// TIA Portal project "Automatizare_RT" (V17) (continued)
REGION Network 14: Cand sistemul hidraulic este in eroare / Wenn das Hydrauliksystem fehlerhaft ist
   RUNG wire#powerrail
      I_Contact( "DB_general".CondOptimePistoane )
      wire#w1
      { S7_GenerateENO := "TRUE" } Move(in := 0, out1 => "DB_Status_Pistoane".Status_Piston_1)
   END_RUNG
   RUNG wire#w1
      { S7_GenerateENO := "TRUE" } Move(in := 0, out1 => "DB_Status_Pistoane".Status_Pison_2)
   END_RUNG
   RUNG wire#w1
      { S7_GenerateENO := "TRUE" } Move(in := 0, out1 => "DB_Status_Pistoane".Status_Piston_A)
   END_RUNG
   RUNG wire#w1
      { S7_GenerateENO := "TRUE" } Move(in := 0, out1 => "DB_Status_Pistoane".Status_Piston_B)
   END_RUNG
   RUNG wire#w1
      { S7_GenerateENO := "TRUE" } Move(in := 0, out1 => "DB_Status_Pistoane".Status_Piston_C)
   END_RUNG
   // the same network as SCL:
   IF NOT "DB_general".CondOptimePistoane THEN
       "DB_Status_Pistoane".Status_Piston_1 := 0;
       "DB_Status_Pistoane".Status_Pison_2 := 0;
       "DB_Status_Pistoane".Status_Piston_A := 0;
       "DB_Status_Pistoane".Status_Piston_B := 0;
       "DB_Status_Pistoane".Status_Piston_C := 0;
   END_IF;
END_REGION
END_FUNCTION

FUNCTION "Status_Motoare" : Void   // FC8, LAD
{ S7_Optimized_Access := 'FALSE' }
VERSION : 0.1
BEGIN

REGION Network 1: motor 1/2 e in functiune
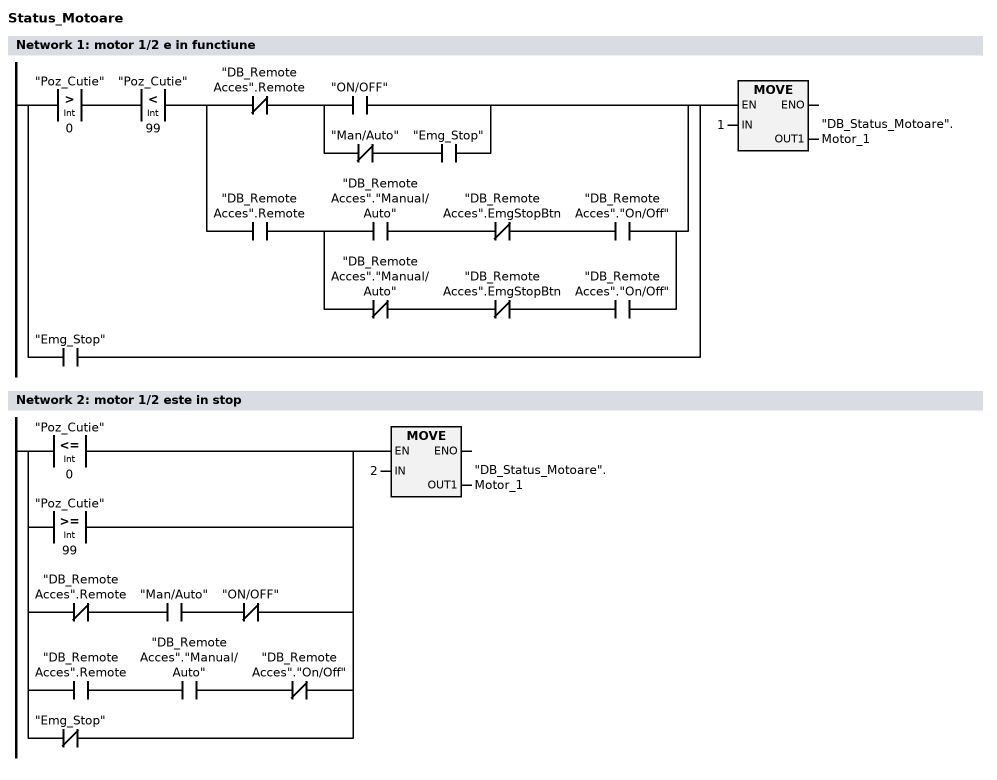
   RUNG wire#powerrail
      { S7_Templates := "SrcType := Int" } GT_Contact(in1 := "Poz_Cutie", in2 := 0)
      { S7_Templates := "SrcType := Int" } LT_Contact(in1 := "Poz_Cutie", in2 := 99)
      wire#w1
      I_Contact( "DB_RemoteAcces".Remote )
      wire#w2
      Contact( "ON/OFF" )
      wire#w3
      { S7_GenerateENO := "TRUE" } Move(in := 1, out1 => "DB_Status_Motoare".Motor_1)
   END_RUNG
   RUNG wire#w2
      I_Contact( "Man/Auto" )
      Contact( "Emg_Stop" )
   END_RUNG wire#w3
   RUNG wire#w1
      Contact( "DB_RemoteAcces".Remote )
      wire#w4
      Contact( "DB_RemoteAcces"."Manual/Auto" )
      I_Contact( "DB_RemoteAcces".EmgStopBtn )
      Contact( "DB_RemoteAcces"."On/Off" )
   END_RUNG wire#w3
   RUNG wire#w4
      I_Contact( "DB_RemoteAcces"."Manual/Auto" )
      I_Contact( "DB_RemoteAcces".EmgStopBtn )
      Contact( "DB_RemoteAcces"."On/Off" )
   END_RUNG wire#w3
   RUNG wire#powerrail
      Contact( "Emg_Stop" )
   END_RUNG wire#w3
   // the same network as SCL:
   IF (("Poz_Cutie" > 0) AND ("Poz_Cutie" < 99) AND ((NOT "DB_RemoteAcces".Remote AND ("ON/OFF" OR (NOT "Man/Auto" AND "Emg_Stop"))) OR ("DB_RemoteAcces".Remote AND (("DB_RemoteAcces"."Manual/Auto" AND NOT "DB_RemoteAcces".EmgStopBtn AND "DB_RemoteAcces"."On/Off") OR (NOT "DB_RemoteAcces"."Manual/Auto" AND NOT "DB_RemoteAcces".EmgStopBtn AND "DB_RemoteAcces"."On/Off"))))) OR "Emg_Stop" THEN
       "DB_Status_Motoare".Motor_1 := 1;
   END_IF;
END_REGION

REGION Network 2: motor 1/2 este in stop
   RUNG wire#powerrail
      { S7_Templates := "SrcType := Int" } LE_Contact(in1 := "Poz_Cutie", in2 := 0)
      wire#w1
      { S7_GenerateENO := "TRUE" } Move(in := 2, out1 => "DB_Status_Motoare".Motor_1)
   END_RUNG
   RUNG wire#powerrail
      { S7_Templates := "SrcType := Int" } GE_Contact(in1 := "Poz_Cutie", in2 := 99)
   END_RUNG wire#w1
   RUNG wire#powerrail
      I_Contact( "DB_RemoteAcces".Remote )
      Contact( "Man/Auto" )
      I_Contact( "ON/OFF" )
   END_RUNG wire#w1
   RUNG wire#powerrail
      Contact( "DB_RemoteAcces".Remote )
      Contact( "DB_RemoteAcces"."Manual/Auto" )
      I_Contact( "DB_RemoteAcces"."On/Off" )
   END_RUNG wire#w1
   RUNG wire#powerrail
      I_Contact( "Emg_Stop" )
   END_RUNG wire#w1
   // the same network as SCL:
   IF ("Poz_Cutie" <= 0) OR ("Poz_Cutie" >= 99) OR (NOT "DB_RemoteAcces".Remote AND "Man/Auto" AND NOT "ON/OFF") OR ("DB_RemoteAcces".Remote AND "DB_RemoteAcces"."Manual/Auto" AND NOT "DB_RemoteAcces"."On/Off") OR NOT "Emg_Stop" THEN
       "DB_Status_Motoare".Motor_1 := 2;
   END_IF;
END_REGION
END_FUNCTION

FUNCTION "CantarFcn" : Void   // FC10, LAD
{ S7_Optimized_Access := 'FALSE' }
VERSION : 0.1
BEGIN

REGION Network 1
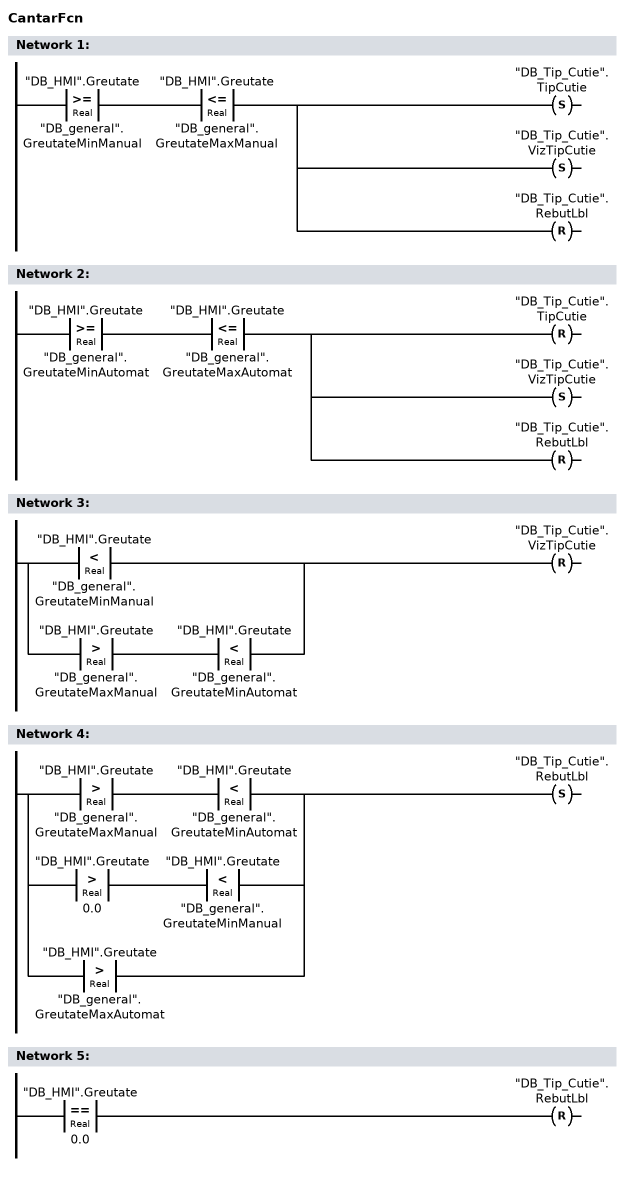
   RUNG wire#powerrail
      { S7_Templates := "SrcType := Real" } GE_Contact(in1 := "DB_HMI".Greutate, in2 := "DB_general".GreutateMinManual)
      { S7_Templates := "SrcType := Real" } LE_Contact(in1 := "DB_HMI".Greutate, in2 := "DB_general".GreutateMaxManual)
      wire#w1
      S_Coil( "DB_Tip_Cutie".TipCutie )
   END_RUNG
   RUNG wire#w1
      S_Coil( "DB_Tip_Cutie".VizTipCutie )
   END_RUNG
   RUNG wire#w1
      R_Coil( "DB_Tip_Cutie".RebutLbl )
   END_RUNG
   // the same network as SCL:
   IF ("DB_HMI".Greutate >= "DB_general".GreutateMinManual) AND ("DB_HMI".Greutate <= "DB_general".GreutateMaxManual) THEN
       "DB_Tip_Cutie".TipCutie := TRUE;
       "DB_Tip_Cutie".VizTipCutie := TRUE;
       "DB_Tip_Cutie".RebutLbl := FALSE;
   END_IF;
END_REGION

REGION Network 2
   RUNG wire#powerrail
      { S7_Templates := "SrcType := Real" } GE_Contact(in1 := "DB_HMI".Greutate, in2 := "DB_general".GreutateMinAutomat)
      { S7_Templates := "SrcType := Real" } LE_Contact(in1 := "DB_HMI".Greutate, in2 := "DB_general".GreutateMaxAutomat)
      wire#w1
      R_Coil( "DB_Tip_Cutie".TipCutie )
   END_RUNG
   RUNG wire#w1
      S_Coil( "DB_Tip_Cutie".VizTipCutie )
   END_RUNG
   RUNG wire#w1
      R_Coil( "DB_Tip_Cutie".RebutLbl )
   END_RUNG
   // the same network as SCL:
   IF ("DB_HMI".Greutate >= "DB_general".GreutateMinAutomat) AND ("DB_HMI".Greutate <= "DB_general".GreutateMaxAutomat) THEN
       "DB_Tip_Cutie".TipCutie := FALSE;
       "DB_Tip_Cutie".VizTipCutie := TRUE;
       "DB_Tip_Cutie".RebutLbl := FALSE;
   END_IF;
END_REGION

REGION Network 3
   RUNG wire#powerrail
      { S7_Templates := "SrcType := Real" } LT_Contact(in1 := "DB_HMI".Greutate, in2 := "DB_general".GreutateMinManual)
      wire#w1
      R_Coil( "DB_Tip_Cutie".VizTipCutie )
   END_RUNG
   RUNG wire#powerrail
      { S7_Templates := "SrcType := Real" } GT_Contact(in1 := "DB_HMI".Greutate, in2 := "DB_general".GreutateMaxManual)
      { S7_Templates := "SrcType := Real" } LT_Contact(in1 := "DB_HMI".Greutate, in2 := "DB_general".GreutateMinAutomat)
   END_RUNG wire#w1
   // the same network as SCL:
   IF ("DB_HMI".Greutate < "DB_general".GreutateMinManual) OR (("DB_HMI".Greutate > "DB_general".GreutateMaxManual) AND ("DB_HMI".Greutate < "DB_general".GreutateMinAutomat)) THEN
       "DB_Tip_Cutie".VizTipCutie := FALSE;
   END_IF;
END_REGION

REGION Network 4
   RUNG wire#powerrail
      { S7_Templates := "SrcType := Real" } GT_Contact(in1 := "DB_HMI".Greutate, in2 := "DB_general".GreutateMaxManual)
      { S7_Templates := "SrcType := Real" } LT_Contact(in1 := "DB_HMI".Greutate, in2 := "DB_general".GreutateMinAutomat)
      wire#w1
      S_Coil( "DB_Tip_Cutie".RebutLbl )
   END_RUNG
   RUNG wire#powerrail
      { S7_Templates := "SrcType := Real" } GT_Contact(in1 := "DB_HMI".Greutate, in2 := 0.0)
      { S7_Templates := "SrcType := Real" } LT_Contact(in1 := "DB_HMI".Greutate, in2 := "DB_general".GreutateMinManual)
   END_RUNG wire#w1
   RUNG wire#powerrail
      { S7_Templates := "SrcType := Real" } GT_Contact(in1 := "DB_HMI".Greutate, in2 := "DB_general".GreutateMaxAutomat)
   END_RUNG wire#w1
   // the same network as SCL:
   IF (("DB_HMI".Greutate > "DB_general".GreutateMaxManual) AND ("DB_HMI".Greutate < "DB_general".GreutateMinAutomat)) OR (("DB_HMI".Greutate > 0.0) AND ("DB_HMI".Greutate < "DB_general".GreutateMinManual)) OR ("DB_HMI".Greutate > "DB_general".GreutateMaxAutomat) THEN
       "DB_Tip_Cutie".RebutLbl := TRUE;
   END_IF;
END_REGION

REGION Network 5
   RUNG wire#powerrail
      { S7_Templates := "SrcType := Real" } EQ_Contact(in1 := "DB_HMI".Greutate, in2 := 0.0)
      R_Coil( "DB_Tip_Cutie".RebutLbl )
   END_RUNG
   // the same network as SCL:
   IF "DB_HMI".Greutate = 0.0 THEN "DB_Tip_Cutie".RebutLbl := FALSE; END_IF;
END_REGION
END_FUNCTION

FUNCTION "CondOptimePistoane" : Void   // FC11, LAD
{ S7_Optimized_Access := 'FALSE' }
VERSION : 0.1
BEGIN

REGION Network 1
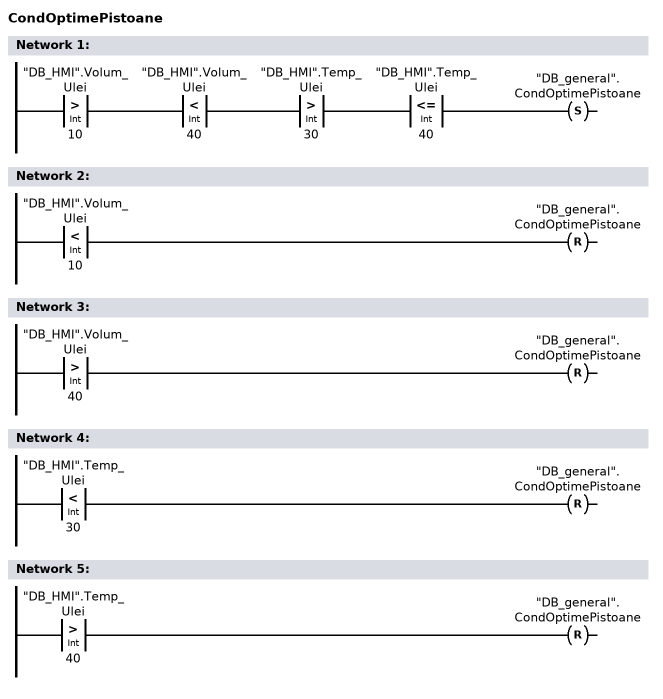
   RUNG wire#powerrail
      { S7_Templates := "SrcType := Int" } GT_Contact(in1 := "DB_HMI".Volum_Ulei, in2 := 10)
      { S7_Templates := "SrcType := Int" } LT_Contact(in1 := "DB_HMI".Volum_Ulei, in2 := 40)
      { S7_Templates := "SrcType := Int" } GT_Contact(in1 := "DB_HMI".Temp_Ulei, in2 := 30)
      { S7_Templates := "SrcType := Int" } LE_Contact(in1 := "DB_HMI".Temp_Ulei, in2 := 40)
      S_Coil( "DB_general".CondOptimePistoane )
   END_RUNG
   // the same network as SCL:
   IF ("DB_HMI".Volum_Ulei > 10) AND ("DB_HMI".Volum_Ulei < 40) AND ("DB_HMI".Temp_Ulei > 30) AND ("DB_HMI".Temp_Ulei <= 40) THEN
       "DB_general".CondOptimePistoane := TRUE;
   END_IF;
END_REGION

REGION Network 2
   RUNG wire#powerrail
      { S7_Templates := "SrcType := Int" } LT_Contact(in1 := "DB_HMI".Volum_Ulei, in2 := 10)
      R_Coil( "DB_general".CondOptimePistoane )
   END_RUNG
   // the same network as SCL:
   IF "DB_HMI".Volum_Ulei < 10 THEN "DB_general".CondOptimePistoane := FALSE; END_IF;
END_REGION

REGION Network 3
   RUNG wire#powerrail
      { S7_Templates := "SrcType := Int" } GT_Contact(in1 := "DB_HMI".Volum_Ulei, in2 := 40)
      R_Coil( "DB_general".CondOptimePistoane )
   END_RUNG
   // the same network as SCL:
   IF "DB_HMI".Volum_Ulei > 40 THEN "DB_general".CondOptimePistoane := FALSE; END_IF;
END_REGION

REGION Network 4
   RUNG wire#powerrail
      { S7_Templates := "SrcType := Int" } LT_Contact(in1 := "DB_HMI".Temp_Ulei, in2 := 30)
      R_Coil( "DB_general".CondOptimePistoane )
   END_RUNG
   // the same network as SCL:
   IF "DB_HMI".Temp_Ulei < 30 THEN "DB_general".CondOptimePistoane := FALSE; END_IF;
END_REGION

REGION Network 5
   RUNG wire#powerrail
      { S7_Templates := "SrcType := Int" } GT_Contact(in1 := "DB_HMI".Temp_Ulei, in2 := 40)
      R_Coil( "DB_general".CondOptimePistoane )
   END_RUNG
   // the same network as SCL:
   IF "DB_HMI".Temp_Ulei > 40 THEN "DB_general".CondOptimePistoane := FALSE; END_IF;
END_REGION
END_FUNCTION

FUNCTION "EroareIntervaleGreutate" : Void   // FC15, STL
{ S7_Optimized_Access := 'FALSE' }
VERSION : 0.1
BEGIN

REGION Network 1


         L     "DB_general".GreutateManual;
         L     "DB_general".Procent_Toleranta;
         *D;
         L     100;
         /R;
         T     "DB_general".TolerantaManual;
         L     "DB_general".TolerantaManual;
         L     "DB_general".GreutateManual;
         +R;
         T     "DB_general".TolerantaManual;
END_REGION
END_FUNCTION

FUNCTION "TipCutieTranzit" : Void   // FC16, LAD
{ S7_Optimized_Access := 'FALSE' }
VERSION : 0.1
BEGIN

REGION Network 1
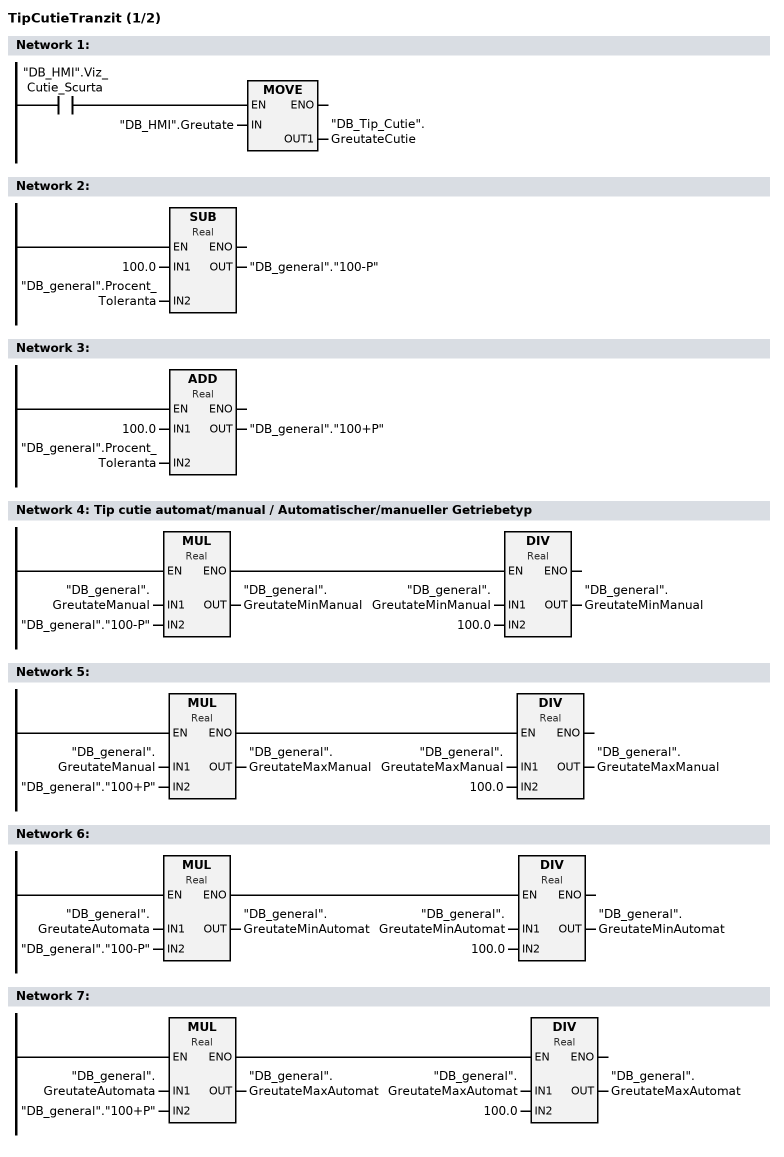
   RUNG wire#powerrail
      Contact( "DB_HMI".Viz_Cutie_Scurta )
      { S7_GenerateENO := "TRUE" } Move(in := "DB_HMI".Greutate, out1 => "DB_Tip_Cutie".GreutateCutie)
   END_RUNG
   // the same network as SCL:
   IF "DB_HMI".Viz_Cutie_Scurta THEN "DB_Tip_Cutie".GreutateCutie := "DB_HMI".Greutate; END_IF;
END_REGION

REGION Network 2
   RUNG wire#powerrail
      { S7_Templates := "SrcType := Real"; S7_GenerateENO := "TRUE" } Sub(in1 := 100.0, in2 := "DB_general".Procent_Toleranta, out => "DB_general"."100-P")
   END_RUNG
   // the same network as SCL:
   "DB_general"."100-P" := 100.0 - "DB_general".Procent_Toleranta;
END_REGION

REGION Network 3
   RUNG wire#powerrail
      { S7_Templates := "SrcType := Real"; S7_GenerateENO := "TRUE" } Add(in1 := 100.0, in2 := "DB_general".Procent_Toleranta, out => "DB_general"."100+P")
   END_RUNG
   // the same network as SCL:
   "DB_general"."100+P" := 100.0 + "DB_general".Procent_Toleranta;
END_REGION

REGION Network 4: Tip cutie automat/manual / Automatischer/manueller Getriebetyp
   RUNG wire#powerrail
      { S7_Templates := "SrcType := Real"; S7_GenerateENO := "TRUE" } Mul(in1 := "DB_general".GreutateManual, in2 := "DB_general"."100-P", out => "DB_general".GreutateMinManual)
      { S7_Templates := "SrcType := Real"; S7_GenerateENO := "TRUE" } Div(in1 := "DB_general".GreutateMinManual, in2 := 100.0, out => "DB_general".GreutateMinManual)
   END_RUNG
   // the same network as SCL:
   // ENO of a box is taken as its EN; it also drops when the box reports an error
   "DB_general".GreutateMinManual := "DB_general".GreutateManual * "DB_general"."100-P";
   "DB_general".GreutateMinManual := "DB_general".GreutateMinManual / 100.0;
END_REGION

REGION Network 5
   RUNG wire#powerrail
      { S7_Templates := "SrcType := Real"; S7_GenerateENO := "TRUE" } Mul(in1 := "DB_general".GreutateManual, in2 := "DB_general"."100+P", out => "DB_general".GreutateMaxManual)
      { S7_Templates := "SrcType := Real"; S7_GenerateENO := "TRUE" } Div(in1 := "DB_general".GreutateMaxManual, in2 := 100.0, out => "DB_general".GreutateMaxManual)
   END_RUNG
   // the same network as SCL:
   // ENO of a box is taken as its EN; it also drops when the box reports an error
   "DB_general".GreutateMaxManual := "DB_general".GreutateManual * "DB_general"."100+P";
   "DB_general".GreutateMaxManual := "DB_general".GreutateMaxManual / 100.0;
END_REGION

REGION Network 6
   RUNG wire#powerrail
      { S7_Templates := "SrcType := Real"; S7_GenerateENO := "TRUE" } Mul(in1 := "DB_general".GreutateAutomata, in2 := "DB_general"."100-P", out => "DB_general".GreutateMinAutomat)
      { S7_Templates := "SrcType := Real"; S7_GenerateENO := "TRUE" } Div(in1 := "DB_general".GreutateMinAutomat, in2 := 100.0, out => "DB_general".GreutateMinAutomat)
   END_RUNG
   // the same network as SCL:
   // ENO of a box is taken as its EN; it also drops when the box reports an error
   "DB_general".GreutateMinAutomat := "DB_general".GreutateAutomata * "DB_general"."100-P";
   "DB_general".GreutateMinAutomat := "DB_general".GreutateMinAutomat / 100.0;
END_REGION

REGION Network 7
   RUNG wire#powerrail
      { S7_Templates := "SrcType := Real"; S7_GenerateENO := "TRUE" } Mul(in1 := "DB_general".GreutateAutomata, in2 := "DB_general"."100+P", out => "DB_general".GreutateMaxAutomat)
      { S7_Templates := "SrcType := Real"; S7_GenerateENO := "TRUE" } Div(in1 := "DB_general".GreutateMaxAutomat, in2 := 100.0, out => "DB_general".GreutateMaxAutomat)
   END_RUNG
   // the same network as SCL:
   // ENO of a box is taken as its EN; it also drops when the box reports an error
   "DB_general".GreutateMaxAutomat := "DB_general".GreutateAutomata * "DB_general"."100+P";
   "DB_general".GreutateMaxAutomat := "DB_general".GreutateMaxAutomat / 100.0;
END_REGION

REGION Network 8
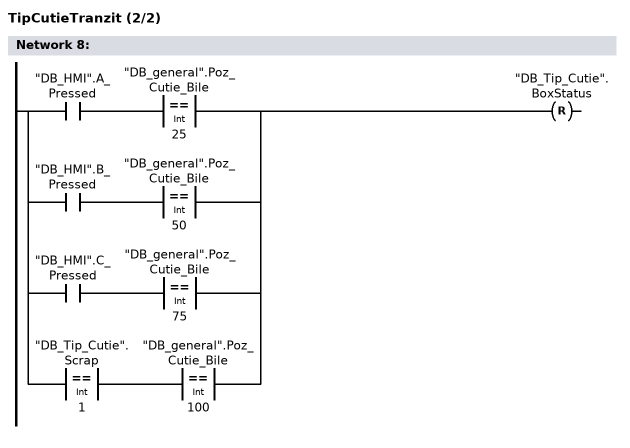
   RUNG wire#powerrail
      Contact( "DB_HMI".A_Pressed )
      { S7_Templates := "SrcType := Int" } EQ_Contact(in1 := "DB_general".Poz_Cutie_Bile, in2 := 25)
      wire#w1
      R_Coil( "DB_Tip_Cutie".BoxStatus )
   END_RUNG
   RUNG wire#powerrail
      Contact( "DB_HMI".B_Pressed )
      { S7_Templates := "SrcType := Int" } EQ_Contact(in1 := "DB_general".Poz_Cutie_Bile, in2 := 50)
   END_RUNG wire#w1
   RUNG wire#powerrail
      Contact( "DB_HMI".C_Pressed )
      { S7_Templates := "SrcType := Int" } EQ_Contact(in1 := "DB_general".Poz_Cutie_Bile, in2 := 75)
   END_RUNG wire#w1
   RUNG wire#powerrail
      { S7_Templates := "SrcType := Int" } EQ_Contact(in1 := "DB_Tip_Cutie".Scrap, in2 := 1)
      { S7_Templates := "SrcType := Int" } EQ_Contact(in1 := "DB_general".Poz_Cutie_Bile, in2 := 100)
   END_RUNG wire#w1
   // the same network as SCL:
   IF ("DB_HMI".A_Pressed AND ("DB_general".Poz_Cutie_Bile = 25)) OR ("DB_HMI".B_Pressed AND ("DB_general".Poz_Cutie_Bile = 50)) OR ("DB_HMI".C_Pressed AND ("DB_general".Poz_Cutie_Bile = 75)) OR (("DB_Tip_Cutie".Scrap = 1) AND ("DB_general".Poz_Cutie_Bile = 100)) THEN
       "DB_Tip_Cutie".BoxStatus := FALSE;
   END_IF;
END_REGION
END_FUNCTION

FUNCTION "EroriCantarire" : Void   // FC17, LAD
{ S7_Optimized_Access := 'FALSE' }
VERSION : 0.1
BEGIN

REGION Network 1
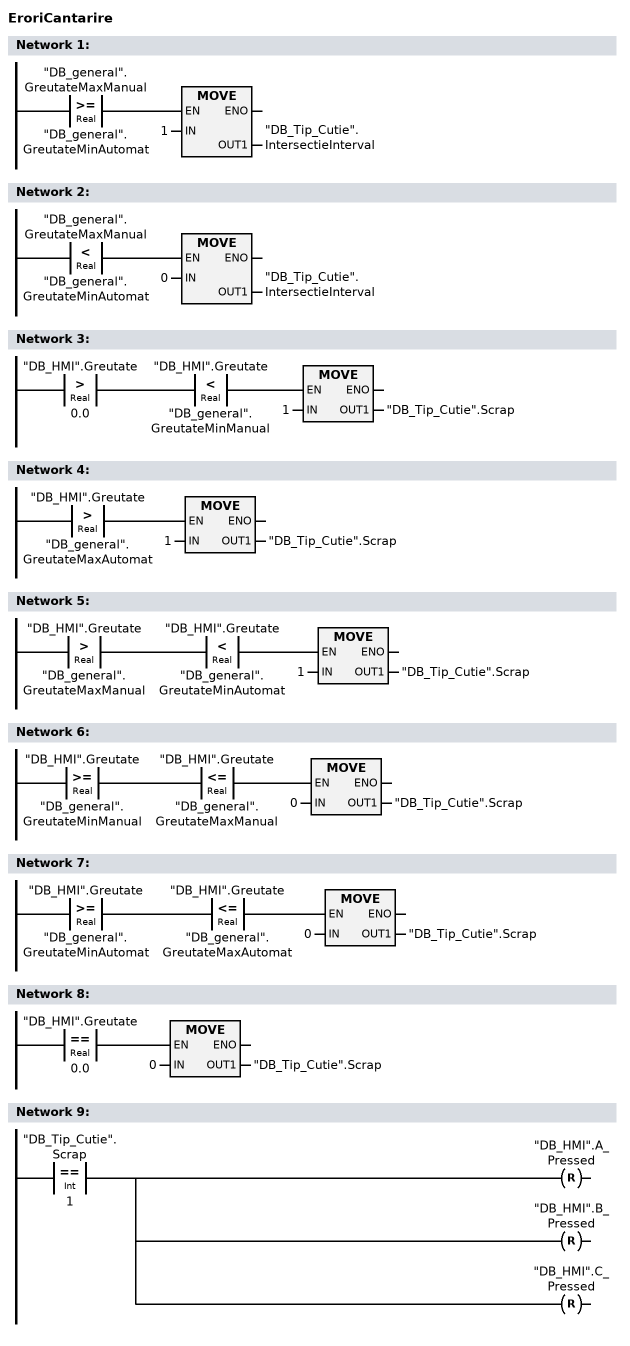
   RUNG wire#powerrail
      { S7_Templates := "SrcType := Real" } GE_Contact(in1 := "DB_general".GreutateMaxManual, in2 := "DB_general".GreutateMinAutomat)
      { S7_GenerateENO := "TRUE" } Move(in := 1, out1 => "DB_Tip_Cutie".IntersectieInterval)
   END_RUNG
   // the same network as SCL:
   IF "DB_general".GreutateMaxManual >= "DB_general".GreutateMinAutomat THEN
       "DB_Tip_Cutie".IntersectieInterval := 1;
   END_IF;
END_REGION

REGION Network 2
   RUNG wire#powerrail
      { S7_Templates := "SrcType := Real" } LT_Contact(in1 := "DB_general".GreutateMaxManual, in2 := "DB_general".GreutateMinAutomat)
      { S7_GenerateENO := "TRUE" } Move(in := 0, out1 => "DB_Tip_Cutie".IntersectieInterval)
   END_RUNG
   // the same network as SCL:
   IF "DB_general".GreutateMaxManual < "DB_general".GreutateMinAutomat THEN
       "DB_Tip_Cutie".IntersectieInterval := 0;
   END_IF;
END_REGION

REGION Network 3
   RUNG wire#powerrail
      { S7_Templates := "SrcType := Real" } GT_Contact(in1 := "DB_HMI".Greutate, in2 := 0.0)
      { S7_Templates := "SrcType := Real" } LT_Contact(in1 := "DB_HMI".Greutate, in2 := "DB_general".GreutateMinManual)
      { S7_GenerateENO := "TRUE" } Move(in := 1, out1 => "DB_Tip_Cutie".Scrap)
   END_RUNG
   // the same network as SCL:
   IF ("DB_HMI".Greutate > 0.0) AND ("DB_HMI".Greutate < "DB_general".GreutateMinManual) THEN
       "DB_Tip_Cutie".Scrap := 1;
   END_IF;
END_REGION

REGION Network 4
   RUNG wire#powerrail
      { S7_Templates := "SrcType := Real" } GT_Contact(in1 := "DB_HMI".Greutate, in2 := "DB_general".GreutateMaxAutomat)
      { S7_GenerateENO := "TRUE" } Move(in := 1, out1 => "DB_Tip_Cutie".Scrap)
   END_RUNG
   // the same network as SCL:
   IF "DB_HMI".Greutate > "DB_general".GreutateMaxAutomat THEN "DB_Tip_Cutie".Scrap := 1; END_IF;
END_REGION

REGION Network 5
   RUNG wire#powerrail
      { S7_Templates := "SrcType := Real" } GT_Contact(in1 := "DB_HMI".Greutate, in2 := "DB_general".GreutateMaxManual)
      { S7_Templates := "SrcType := Real" } LT_Contact(in1 := "DB_HMI".Greutate, in2 := "DB_general".GreutateMinAutomat)
      { S7_GenerateENO := "TRUE" } Move(in := 1, out1 => "DB_Tip_Cutie".Scrap)
   END_RUNG
   // the same network as SCL:
   IF ("DB_HMI".Greutate > "DB_general".GreutateMaxManual) AND ("DB_HMI".Greutate < "DB_general".GreutateMinAutomat) THEN
       "DB_Tip_Cutie".Scrap := 1;
   END_IF;
END_REGION

REGION Network 6
   RUNG wire#powerrail
      { S7_Templates := "SrcType := Real" } GE_Contact(in1 := "DB_HMI".Greutate, in2 := "DB_general".GreutateMinManual)
      { S7_Templates := "SrcType := Real" } LE_Contact(in1 := "DB_HMI".Greutate, in2 := "DB_general".GreutateMaxManual)
      { S7_GenerateENO := "TRUE" } Move(in := 0, out1 => "DB_Tip_Cutie".Scrap)
   END_RUNG
   // the same network as SCL:
   IF ("DB_HMI".Greutate >= "DB_general".GreutateMinManual) AND ("DB_HMI".Greutate <= "DB_general".GreutateMaxManual) THEN
       "DB_Tip_Cutie".Scrap := 0;
   END_IF;
END_REGION

REGION Network 7
   RUNG wire#powerrail
      { S7_Templates := "SrcType := Real" } GE_Contact(in1 := "DB_HMI".Greutate, in2 := "DB_general".GreutateMinAutomat)
      { S7_Templates := "SrcType := Real" } LE_Contact(in1 := "DB_HMI".Greutate, in2 := "DB_general".GreutateMaxAutomat)
      { S7_GenerateENO := "TRUE" } Move(in := 0, out1 => "DB_Tip_Cutie".Scrap)
   END_RUNG
   // the same network as SCL:
   IF ("DB_HMI".Greutate >= "DB_general".GreutateMinAutomat) AND ("DB_HMI".Greutate <= "DB_general".GreutateMaxAutomat) THEN
       "DB_Tip_Cutie".Scrap := 0;
   END_IF;
END_REGION

REGION Network 8
   RUNG wire#powerrail
      { S7_Templates := "SrcType := Real" } EQ_Contact(in1 := "DB_HMI".Greutate, in2 := 0.0)
      { S7_GenerateENO := "TRUE" } Move(in := 0, out1 => "DB_Tip_Cutie".Scrap)
   END_RUNG
   // the same network as SCL:
   IF "DB_HMI".Greutate = 0.0 THEN "DB_Tip_Cutie".Scrap := 0; END_IF;
END_REGION

REGION Network 9
   RUNG wire#powerrail
      { S7_Templates := "SrcType := Int" } EQ_Contact(in1 := "DB_Tip_Cutie".Scrap, in2 := 1)
      wire#w1
      R_Coil( "DB_HMI".A_Pressed )
   END_RUNG
   RUNG wire#w1
      R_Coil( "DB_HMI".B_Pressed )
   END_RUNG
   RUNG wire#w1
      R_Coil( "DB_HMI".C_Pressed )
   END_RUNG
   // the same network as SCL:
   IF "DB_Tip_Cutie".Scrap = 1 THEN
       "DB_HMI".A_Pressed := FALSE;
       "DB_HMI".B_Pressed := FALSE;
       "DB_HMI".C_Pressed := FALSE;
   END_IF;
END_REGION
END_FUNCTION

FUNCTION "ConsolaComanda" : Void   // FC21, LAD
{ S7_Optimized_Access := 'FALSE' }
VERSION : 0.1
   VAR_TEMP   // added for the SCL form of the ladder/FBD networks
      _w1 : Bool;
   END_VAR
BEGIN

REGION Network 1
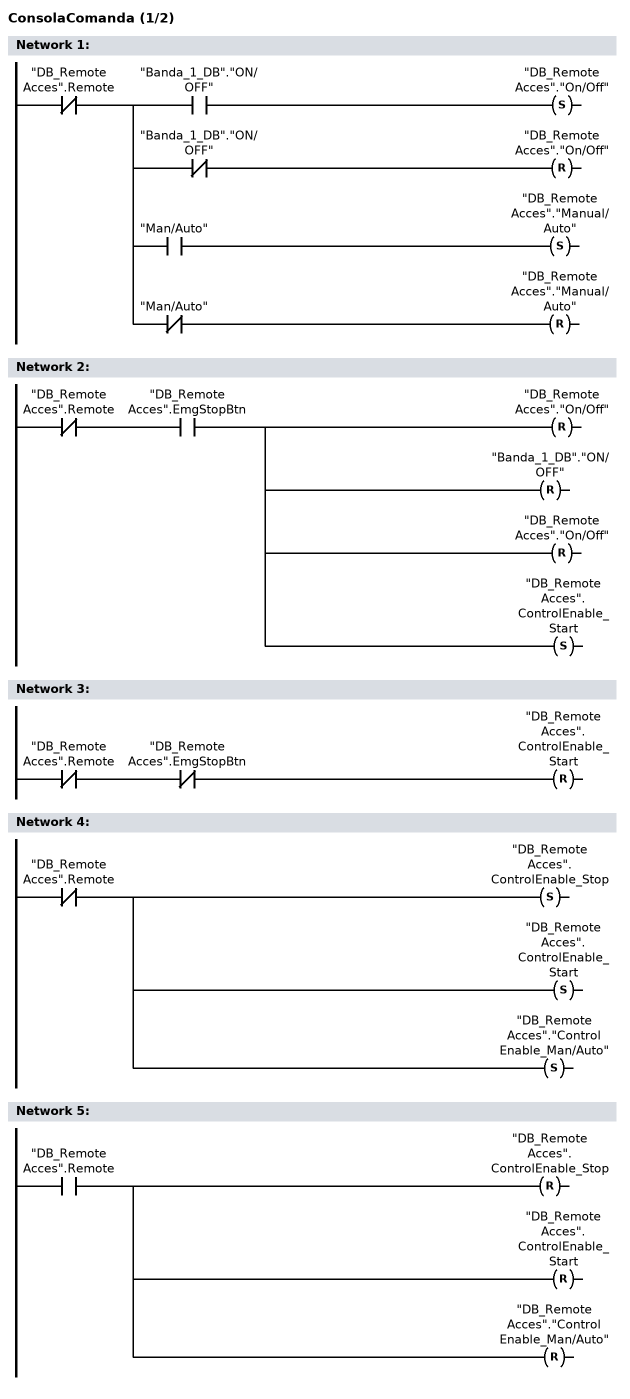
   RUNG wire#powerrail
      I_Contact( "DB_RemoteAcces".Remote )
      wire#w1
      Contact( "Banda_1_DB"."ON/OFF" )
      S_Coil( "DB_RemoteAcces"."On/Off" )
   END_RUNG
   RUNG wire#w1
      I_Contact( "Banda_1_DB"."ON/OFF" )
      R_Coil( "DB_RemoteAcces"."On/Off" )
   END_RUNG
   RUNG wire#w1
      Contact( "Man/Auto" )
      S_Coil( "DB_RemoteAcces"."Manual/Auto" )
   END_RUNG
   RUNG wire#w1
      I_Contact( "Man/Auto" )
      R_Coil( "DB_RemoteAcces"."Manual/Auto" )
   END_RUNG
   // the same network as SCL:
   #_w1 := NOT "DB_RemoteAcces".Remote;
   IF #_w1 AND "Banda_1_DB"."ON/OFF" THEN "DB_RemoteAcces"."On/Off" := TRUE; END_IF;
   IF #_w1 AND NOT "Banda_1_DB"."ON/OFF" THEN "DB_RemoteAcces"."On/Off" := FALSE; END_IF;
   IF #_w1 AND "Man/Auto" THEN "DB_RemoteAcces"."Manual/Auto" := TRUE; END_IF;
   IF #_w1 AND NOT "Man/Auto" THEN "DB_RemoteAcces"."Manual/Auto" := FALSE; END_IF;
END_REGION

REGION Network 2
   RUNG wire#powerrail
      I_Contact( "DB_RemoteAcces".Remote )
      Contact( "DB_RemoteAcces".EmgStopBtn )
      wire#w1
      R_Coil( "DB_RemoteAcces"."On/Off" )
   END_RUNG
   RUNG wire#w1
      R_Coil( "Banda_1_DB"."ON/OFF" )
   END_RUNG
   RUNG wire#w1
      R_Coil( "DB_RemoteAcces"."On/Off" )
   END_RUNG
   RUNG wire#w1
      S_Coil( "DB_RemoteAcces".ControlEnable_Start )
   END_RUNG
   // the same network as SCL:
   IF NOT "DB_RemoteAcces".Remote AND "DB_RemoteAcces".EmgStopBtn THEN
       "DB_RemoteAcces"."On/Off" := FALSE;
       "Banda_1_DB"."ON/OFF" := FALSE;
       "DB_RemoteAcces"."On/Off" := FALSE;
       "DB_RemoteAcces".ControlEnable_Start := TRUE;
   END_IF;
END_REGION

REGION Network 3
   RUNG wire#powerrail
      I_Contact( "DB_RemoteAcces".Remote )
      I_Contact( "DB_RemoteAcces".EmgStopBtn )
      R_Coil( "DB_RemoteAcces".ControlEnable_Start )
   END_RUNG
   // the same network as SCL:
   IF NOT "DB_RemoteAcces".Remote AND NOT "DB_RemoteAcces".EmgStopBtn THEN
       "DB_RemoteAcces".ControlEnable_Start := FALSE;
   END_IF;
END_REGION

REGION Network 4
   RUNG wire#powerrail
      I_Contact( "DB_RemoteAcces".Remote )
      wire#w1
      S_Coil( "DB_RemoteAcces".ControlEnable_Stop )
   END_RUNG
   RUNG wire#w1
      S_Coil( "DB_RemoteAcces".ControlEnable_Start )
   END_RUNG
   RUNG wire#w1
      S_Coil( "DB_RemoteAcces"."ControlEnable_Man/Auto" )
   END_RUNG
   // the same network as SCL:
   IF NOT "DB_RemoteAcces".Remote THEN
       "DB_RemoteAcces".ControlEnable_Stop := TRUE;
       "DB_RemoteAcces".ControlEnable_Start := TRUE;
       "DB_RemoteAcces"."ControlEnable_Man/Auto" := TRUE;
   END_IF;
END_REGION

REGION Network 5
   RUNG wire#powerrail
      Contact( "DB_RemoteAcces".Remote )
      wire#w1
      R_Coil( "DB_RemoteAcces".ControlEnable_Stop )
   END_RUNG
   RUNG wire#w1
      R_Coil( "DB_RemoteAcces".ControlEnable_Start )
   END_RUNG
   RUNG wire#w1
      R_Coil( "DB_RemoteAcces"."ControlEnable_Man/Auto" )
   END_RUNG
   // the same network as SCL:
   IF "DB_RemoteAcces".Remote THEN
       "DB_RemoteAcces".ControlEnable_Stop := FALSE;
       "DB_RemoteAcces".ControlEnable_Start := FALSE;
       "DB_RemoteAcces"."ControlEnable_Man/Auto" := FALSE;
   END_IF;
END_REGION

REGION Network 6
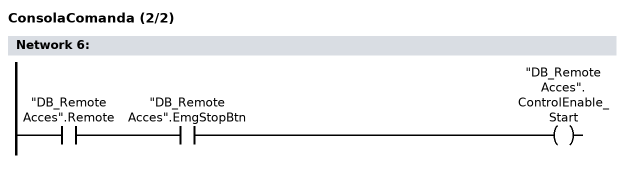
   RUNG wire#powerrail
      Contact( "DB_RemoteAcces".Remote )
      Contact( "DB_RemoteAcces".EmgStopBtn )
      Coil( "DB_RemoteAcces".ControlEnable_Start )
   END_RUNG
   // the same network as SCL:
   "DB_RemoteAcces".ControlEnable_Start := "DB_RemoteAcces".Remote AND "DB_RemoteAcces".EmgStopBtn;
END_REGION
END_FUNCTION

// folder: Hidraulic/Functii

FUNCTION "Adaugare/Scadere_Ulei" : Void   // FC2, LAD
{ S7_Optimized_Access := 'FALSE' }
VERSION : 0.1
BEGIN

REGION Network 1
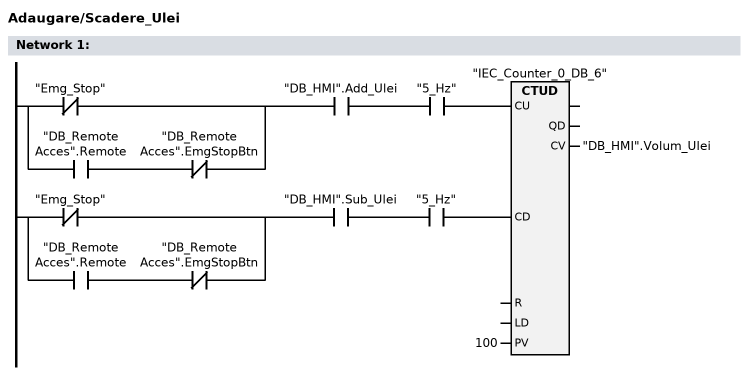
   "IEC_Counter_0_DB_6".CTUD(CU := (NOT "Emg_Stop" OR ("DB_RemoteAcces".Remote AND NOT "DB_RemoteAcces".EmgStopBtn)) AND "DB_HMI".Add_Ulei AND "5_Hz",
                           CD := (NOT "Emg_Stop" OR ("DB_RemoteAcces".Remote AND NOT "DB_RemoteAcces".EmgStopBtn)) AND "DB_HMI".Sub_Ulei AND "5_Hz",
                           PV := 100,
                           CV => "DB_HMI".Volum_Ulei);
END_REGION
END_FUNCTION

FUNCTION "Temp_Ulei" : Void   // FC3, LAD
{ S7_Optimized_Access := 'FALSE' }
VERSION : 0.1
BEGIN

REGION Network 1
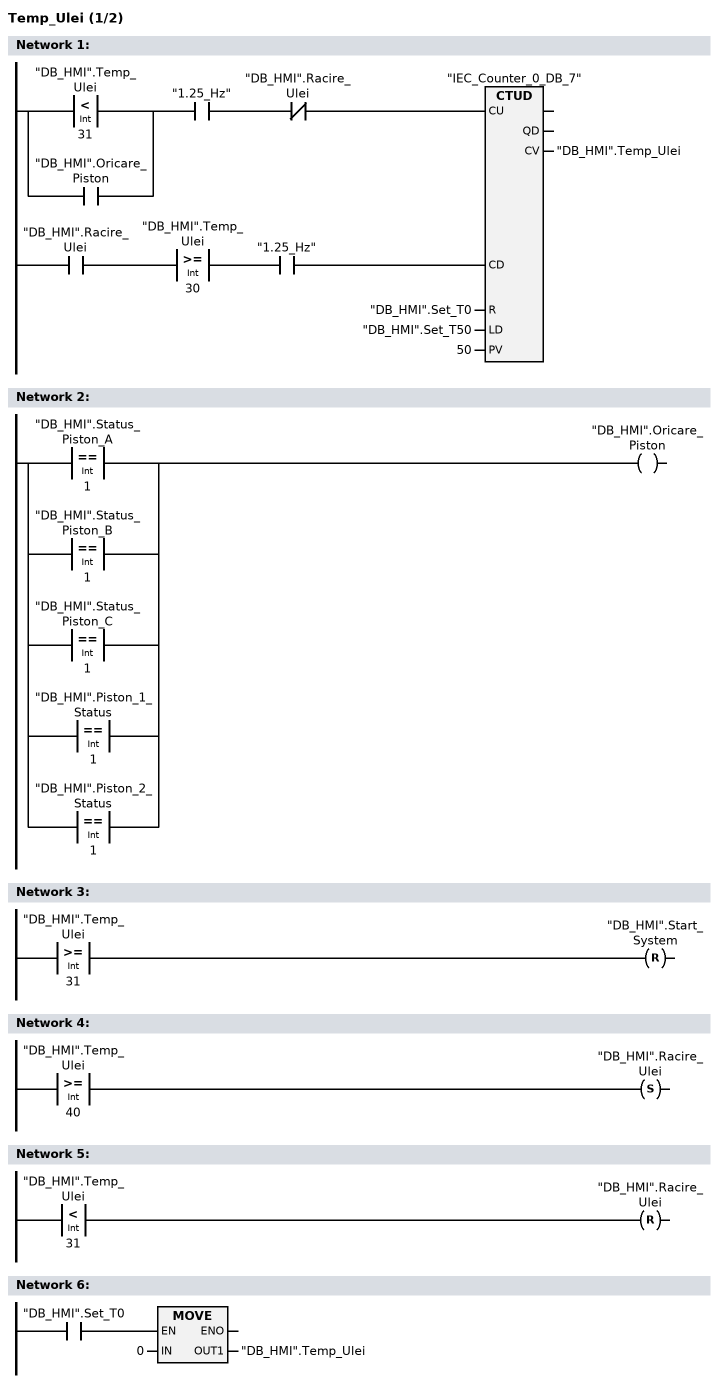
   "IEC_Counter_0_DB_7".CTUD(CU := (("DB_HMI".Temp_Ulei < 31) OR "DB_HMI".Oricare_Piston) AND "1.25_Hz" AND NOT "DB_HMI".Racire_Ulei,
                           CD := "DB_HMI".Racire_Ulei AND ("DB_HMI".Temp_Ulei >= 30) AND "1.25_Hz",
                           R := "DB_HMI".Set_T0,
                           LD := "DB_HMI".Set_T50,
                           PV := 50,
                           CV => "DB_HMI".Temp_Ulei);
END_REGION

REGION Network 2
   RUNG wire#powerrail
      { S7_Templates := "SrcType := Int" } EQ_Contact(in1 := "DB_HMI".Status_Piston_A, in2 := 1)
      wire#w1
      Coil( "DB_HMI".Oricare_Piston )
   END_RUNG
   RUNG wire#powerrail
      { S7_Templates := "SrcType := Int" } EQ_Contact(in1 := "DB_HMI".Status_Piston_B, in2 := 1)
   END_RUNG wire#w1
   RUNG wire#powerrail
      { S7_Templates := "SrcType := Int" } EQ_Contact(in1 := "DB_HMI".Status_Piston_C, in2 := 1)
   END_RUNG wire#w1
   RUNG wire#powerrail
      { S7_Templates := "SrcType := Int" } EQ_Contact(in1 := "DB_HMI".Piston_1_Status, in2 := 1)
   END_RUNG wire#w1
   RUNG wire#powerrail
      { S7_Templates := "SrcType := Int" } EQ_Contact(in1 := "DB_HMI".Piston_2_Status, in2 := 1)
   END_RUNG wire#w1
   // the same network as SCL:
   "DB_HMI".Oricare_Piston := ("DB_HMI".Status_Piston_A = 1) OR ("DB_HMI".Status_Piston_B = 1) OR ("DB_HMI".Status_Piston_C = 1) OR ("DB_HMI".Piston_1_Status = 1) OR ("DB_HMI".Piston_2_Status = 1);
END_REGION

REGION Network 3
   RUNG wire#powerrail
      { S7_Templates := "SrcType := Int" } GE_Contact(in1 := "DB_HMI".Temp_Ulei, in2 := 31)
      R_Coil( "DB_HMI".Start_System )
   END_RUNG
   // the same network as SCL:
   IF "DB_HMI".Temp_Ulei >= 31 THEN "DB_HMI".Start_System := FALSE; END_IF;
END_REGION

REGION Network 4
   RUNG wire#powerrail
      { S7_Templates := "SrcType := Int" } GE_Contact(in1 := "DB_HMI".Temp_Ulei, in2 := 40)
      S_Coil( "DB_HMI".Racire_Ulei )
   END_RUNG
   // the same network as SCL:
   IF "DB_HMI".Temp_Ulei >= 40 THEN "DB_HMI".Racire_Ulei := TRUE; END_IF;
END_REGION

REGION Network 5
   RUNG wire#powerrail
      { S7_Templates := "SrcType := Int" } LT_Contact(in1 := "DB_HMI".Temp_Ulei, in2 := 31)
      R_Coil( "DB_HMI".Racire_Ulei )
   END_RUNG
   // the same network as SCL:
   IF "DB_HMI".Temp_Ulei < 31 THEN "DB_HMI".Racire_Ulei := FALSE; END_IF;
END_REGION

REGION Network 6
   RUNG wire#powerrail
      Contact( "DB_HMI".Set_T0 )
      { S7_GenerateENO := "TRUE" } Move(in := 0, out1 => "DB_HMI".Temp_Ulei)
   END_RUNG
   // the same network as SCL:
   IF "DB_HMI".Set_T0 THEN "DB_HMI".Temp_Ulei := 0; END_IF;
END_REGION

REGION Network 7: pompeaza aer cald / pumpt heiße LufT
